      { S7_Templates := "SrcType := Real" } EQ_Contact(in1 := "MB_MFC_FLOAT_DB".FCounterLimit, in2 := "MB_MFC_FLOAT_DB".MFC401_VOL_SP)
      { S7_Templates := "SrcType := Real" } LT_Contact(in1 := "PT402_VAL", in2 := "PT402_HIGH")
      { S7_Templates := "SrcType := Real" } GE_Contact(in1 := "PT601_VAL", in2 := "PT401_CALC_50PRCT")
      wire#w9
      I_Contact( "S6_3" )
      wire#w10
      Coil( "S6_2" )
   END_RUNG
   RUNG wire#w8
      Contact( "S6_2" )
   END_RUNG wire#w9
   RUNG wire#w10
      Move(in := -1, out1 => "MB_MFC_FLOAT_DB"."STEP")
      Move(in := 0, out1 => "MB_MFC_INT_DB".MFC_Setpoint)
      Move(in := 40, out1 => "MB_MFC_INT_DB".START_STEP)   // Closes Valve
      S_Coil( "MB_MFC_INT_DB".LOAD_STEP )
   END_RUNG
   RUNG wire#w10
      S_Coil( "PV702_NC" )
   END_RUNG
   RUNG wire#powerrail
      Contact( #RUN )
      wire#w11
      Contact( "S6_2" )
      I_Contact( "PV702_NOT_OPEN_LS" )
      wire#w12
      { S7_Templates := "SrcType := SInt" } GE_Contact(in1 := "MB_MFC_INT_DB"."STEP", in2 := 2)
      { S7_Templates := "SrcType := UInt" } EQ_Contact(in1 := "MB_MFC_INT_DB".ControlMode, in2 := 0)
      { S7_Templates := "SrcType := UInt" } EQ_Contact(in1 := "MB_MFC_INT_DB".ValveOutput, in2 := 0)
      { S7_Templates := "SrcType := UInt" } EQ_Contact(in1 := "MB_MFC_INT_DB".Measure, in2 := 0)
      wire#w13
      I_Contact( "S6_3A" )
      wire#w14
      Coil( "S6_3" )
   END_RUNG
   RUNG wire#w12
      { S7_Templates := "SrcType := Real" } LE_Contact(in1 := "PT601_VAL", in2 := "PT901_VAL")
   END_RUNG wire#w13
   RUNG wire#w11
      Contact( "S6_3" )
   END_RUNG wire#w13
   RUNG wire#w14
      R_Coil( "PV702_NC" )
   END_RUNG
   RUNG wire#powerrail
      Contact( #RUN )
      wire#w15
      Contact( "S6_3" )
      I_Contact( "PV702_NOT_CLOSED_LS" )
      { S7_Templates := "SrcType := SInt" } GE_Contact(in1 := "MB_MFC_INT_DB"."STEP", in2 := 3)
      { S7_Templates := "SrcType := UInt" } EQ_Contact(in1 := "MB_MFC_INT_DB".CounterMode, in2 := 2)
      { S7_Templates := "SrcType := UInt" } EQ_Contact(in1 := "MB_MFC_INT_DB".CounterVal, in2 := 0)
      { S7_Templates := "SrcType := UInt" } EQ_Contact(in1 := "MB_MFC_INT_DB".ValveOutput, in2 := 0)
      { S7_Templates := "SrcType := UInt" } EQ_Contact(in1 := "MB_MFC_INT_DB".Measure, in2 := 0)
      I_Contact( #ALARM )
      wire#w16
      I_Contact( "S6_3B" )
      wire#w17
      Coil( "S6_3A" )
   END_RUNG
   RUNG wire#w15
      Contact( "S6_3A" )
   END_RUNG wire#w16
   RUNG wire#w17
      Move(in := -1, out1 => "MB_MFC_INT_DB"."STEP")
      Move(in := -1, out1 => "MB_MFC_FLOAT_DB"."STEP")
   END_RUNG
   RUNG wire#powerrail
      Contact( #RUN )
      wire#w18
      Contact( "S6_3A" )
      Contact( "IEC_Timer_S6_DB_1".Q )
      I_Contact( #ALARM )
      wire#w19
      I_Contact( "S6_4" )
      wire#w20
      Coil( "S6_3B" )
   END_RUNG
   RUNG wire#w18
      Contact( "S6_3B" )
   END_RUNG wire#w19
   RUNG wire#w20
      S_Coil( "PV701_NC" )
   END_RUNG
   RUNG wire#w20
      Move(in := "MB_MFC_FLOAT_DB".MFC401_FLOW_SP, out1 => "MB_MFC_FLOAT_DB".FLOW_SP)
      Move(in := 20, out1 => "MB_MFC_FLOAT_DB".START_STEP)
      S_Coil( "MB_MFC_FLOAT_DB".LOAD_STEP )
   END_RUNG
   RUNG wire#powerrail
      Contact( #RUN )
      wire#w21
      Contact( "S6_3B" )
      I_Contact( "PV701_NOT_OPEN_LS" )
      { S7_Templates := "SrcType := SInt" } EQ_Contact(in1 := "MB_MFC_FLOAT_DB"."STEP", in2 := 2)
      wire#w22
      I_Contact( "S6_5" )
      wire#w23
      Coil( "S6_4" )
   END_RUNG
   RUNG wire#w21
      Contact( "S6_4" )
   END_RUNG wire#w22
   RUNG wire#w23
      Move(in := -1, out1 => "MB_MFC_INT_DB"."STEP")
   END_RUNG
   RUNG wire#powerrail
      Contact( #RUN )
      wire#w24
      Contact( "S6_4" )
      wire#w25
      { S7_Templates := "SrcType := SInt" } GE_Contact(in1 := "MB_MFC_FLOAT_DB"."STEP", in2 := 1)
      { S7_Templates := "SrcType := Real" } GE_Contact(in1 := "MB_MFC_FLOAT_DB".FCounterVal, in2 := "MB_MFC_FLOAT_DB".COUNTER_LIMIT_SP)
      wire#w26
      I_Contact( "S6_6" )
      wire#w27
      Coil( "S6_5" )
   END_RUNG
   RUNG wire#w25
      { S7_Templates := "SrcType := Real" } GE_Contact(in1 := "PT901_VAL", in2 := "PT901_SP_H")
   END_RUNG wire#w26
   RUNG wire#w24
      Contact( "S6_5" )
   END_RUNG wire#w26
   RUNG wire#w27
      R_Coil( "PV401_NC" )
      R_Coil( "PV701_NC" )
   END_RUNG
   RUNG wire#w27
      Move(in := -1, out1 => "MB_MFC_FLOAT_DB"."STEP")
      Move(in := "MFC_601_MB_ADDR", out1 => "MB_MFC_INT_DB".MFC_ADDRESS)
      Move(in := 68, out1 => "MB_MFC_INT_DB".START_STEP)   // Purge Valve
      S_Coil( "MB_MFC_INT_DB".LOAD_STEP )
   END_RUNG
   RUNG wire#powerrail
      Contact( #RUN )
      wire#w28
      Contact( "S6_5" )
      I_Contact( "PV701_NOT_CLOSED_LS" )
      { S7_Templates := "SrcType := UInt" } EQ_Contact(in1 := "MB_MFC_INT_DB".ControlMode, in2 := 8)
      { S7_Templates := "SrcType := SInt" } EQ_Contact(in1 := "MB_MFC_INT_DB"."STEP", in2 := 4)
      wire#w29
      I_Contact( "S6_7" )
      wire#w30
      Coil( "S6_6" )
   END_RUNG
   RUNG wire#w28
      Contact( "S6_6" )
   END_RUNG wire#w29
   RUNG wire#w30
      S_Coil( "PV702_NC" )
   END_RUNG
   RUNG wire#w30
      Move(in := -1, out1 => "MB_MFC_INT_DB"."STEP")
   END_RUNG
   RUNG wire#powerrail
      Contact( #RUN )
      wire#w31
      Contact( "S6_6" )
      I_Contact( "PV702_NOT_OPEN_LS" )
      { S7_Templates := "SrcType := Real" } LE_Contact(in1 := "PT601_VAL", in2 := "PT601_ZERO")
      wire#w32
      I_Contact( "S6_8" )
      wire#w33
      Coil( "S6_7" )
   END_RUNG
   RUNG wire#w31
      Contact( "S6_7" )
   END_RUNG wire#w32
   RUNG wire#w33
      R_Coil( "PV602_NC" )
      R_Coil( "PV402_NC" )
   END_RUNG
   RUNG wire#w33
      R_Coil( "PV702_NC" )
   END_RUNG
   RUNG wire#w33
      Move(in := "MFC_601_MB_ADDR", out1 => "MB_MFC_INT_DB".MFC_ADDRESS)
      Move(in := "MB_VAL_CONTROL_MODE_BUS", out1 => "MB_MFC_INT_DB".MFC_MODE_SP)
      Move(in := 0, out1 => "MB_MFC_INT_DB".MFC_Setpoint)
      Move(in := 10, out1 => "MB_MFC_INT_DB".START_STEP)
      S_Coil( "MB_MFC_INT_DB".LOAD_STEP )
   END_RUNG
   RUNG wire#powerrail
      Contact( #RUN )
      wire#w34
      Contact( "S6_7" )
      I_Contact( "PV702_NOT_CLOSED_LS" )
      { S7_Templates := "SrcType := SInt" } EQ_Contact(in1 := "MB_MFC_INT_DB"."STEP", in2 := 4)
      { S7_Templates := "SrcType := UInt" } EQ_Contact(in1 := "MB_MFC_INT_DB".ControlMode, in2 := 0)
      Contact( "IEC_Timer_S6_DB_1".Q )
      wire#w35
      I_Contact( "S6_9" )
      wire#w36
      Coil( "S6_8" )
   END_RUNG
   RUNG wire#w34
      Contact( "S6_8" )
   END_RUNG wire#w35
   RUNG wire#w36
      R_Coil( "PV403_NO" )
   END_RUNG
   RUNG wire#w36
      { S7_GenerateENO := "TRUE" } Move(in := "PT901_VAL", out1 => "PT901_END_H")
   END_RUNG
   RUNG wire#w36
      Contact( "AlwaysFALSE" )
      Move(in := -1, out1 => "MB_MFC_INT_DB"."STEP")
      Move(in := -1, out1 => "MB_MFC_FLOAT_DB"."STEP")
   END_RUNG
   RUNG wire#powerrail
      Contact( #RUN )
      wire#w37
      Contact( "S6_8" )
      { S7_Templates := "SrcType := Real" } LE_Contact(in1 := "PT402_VAL", in2 := 0.0)
      wire#w38
      Coil( "S6_9" )
   END_RUNG
   RUNG wire#w37
      Contact( "S6_9" )
   END_RUNG wire#w38
   RUNG wire#w38
      Coil( #ENDED )
   END_RUNG
   // the same network as SCL:
   #_w1 := #RUN AND "AUTO_CYCLE" AND #RUN AND NOT "S6_M";   // rising edge of #RUN
   "S6_M" := #RUN;
   "S6_0" := ((((#RUN AND #START) OR #_w1) AND NOT #ALARM) OR (#RUN AND "S6_0")) AND NOT "S6_1";
   IF "S6_0" THEN
       "MB_MFC_FLOAT_DB".MFC_ADDRESS := "MFC_401_MB_ADDR";
       "MB_MFC_FLOAT_DB"."STEP" := -1;
       "MB_MFC_INT_DB".MFC_MODE_SP := "MB_VAL_CONTROL_MODE_BUS";
       "MB_MFC_INT_DB".START_STEP := 10;
       "MB_MFC_INT_DB".LOAD_STEP := TRUE;
       "MB_MFC_INT_DB".MFC_ADDRESS := "MFC_401_MB_ADDR";
       "GREEN_LIGHT" := FALSE;
       "YELLOW_LIGHT" := FALSE;
       "RED_ON" := TRUE;
   END_IF;
   "S6_1" := #RUN AND (("S6_0" AND "IEC_Timer_S6_DB_1".Q AND NOT #ALARM) OR "S6_1") AND NOT "S6_2";
   IF "S6_1" THEN
       "PV403_NO" := TRUE;
       "PV401_NC" := TRUE;
       "PV402_NC" := TRUE;
       "PV602_NC" := TRUE;
       "MB_MFC_INT_DB"."STEP" := -1;
       "MB_MFC_FLOAT_DB".FLOW_SP := 2.0;
       "MB_MFC_FLOAT_DB".START_STEP := 20;
       "MB_MFC_FLOAT_DB".LOAD_STEP := TRUE;
   END_IF;
   "S6_2" := #RUN AND (("S6_1" AND ("MB_MFC_FLOAT_DB"."STEP" >= 4) AND ("MB_MFC_FLOAT_DB".FCounterLimit = "MB_MFC_FLOAT_DB".MFC401_VOL_SP) AND ("PT402_VAL" < "PT402_HIGH") AND ("PT601_VAL" >= "PT401_CALC_50PRCT")) OR "S6_2") AND NOT "S6_3";
   IF "S6_2" THEN
       "MB_MFC_FLOAT_DB"."STEP" := -1;
       "MB_MFC_INT_DB".MFC_Setpoint := 0;
       "MB_MFC_INT_DB".START_STEP := 40;   // Closes Valve
       "MB_MFC_INT_DB".LOAD_STEP := TRUE;
       "PV702_NC" := TRUE;
   END_IF;
   "S6_3" := #RUN AND (("S6_2" AND NOT "PV702_NOT_OPEN_LS" AND ((("MB_MFC_INT_DB"."STEP" >= 2) AND ("MB_MFC_INT_DB".ControlMode = 0) AND ("MB_MFC_INT_DB".ValveOutput = 0) AND ("MB_MFC_INT_DB".Measure = 0)) OR ("PT601_VAL" <= "PT901_VAL"))) OR "S6_3") AND NOT "S6_3A";
   IF "S6_3" THEN "PV702_NC" := FALSE; END_IF;
   "S6_3A" := #RUN AND (("S6_3" AND NOT "PV702_NOT_CLOSED_LS" AND ("MB_MFC_INT_DB"."STEP" >= 3) AND ("MB_MFC_INT_DB".CounterMode = 2) AND ("MB_MFC_INT_DB".CounterVal = 0) AND ("MB_MFC_INT_DB".ValveOutput = 0) AND ("MB_MFC_INT_DB".Measure = 0) AND NOT #ALARM) OR "S6_3A") AND NOT "S6_3B";
   IF "S6_3A" THEN
       "MB_MFC_INT_DB"."STEP" := -1;
       "MB_MFC_FLOAT_DB"."STEP" := -1;
   END_IF;
   "S6_3B" := #RUN AND (("S6_3A" AND "IEC_Timer_S6_DB_1".Q AND NOT #ALARM) OR "S6_3B") AND NOT "S6_4";
   IF "S6_3B" THEN
       "PV701_NC" := TRUE;
       "MB_MFC_FLOAT_DB".FLOW_SP := "MB_MFC_FLOAT_DB".MFC401_FLOW_SP;
       "MB_MFC_FLOAT_DB".START_STEP := 20;
       "MB_MFC_FLOAT_DB".LOAD_STEP := TRUE;
   END_IF;
   "S6_4" := #RUN AND (("S6_3B" AND NOT "PV701_NOT_OPEN_LS" AND ("MB_MFC_FLOAT_DB"."STEP" = 2)) OR "S6_4") AND NOT "S6_5";
   IF "S6_4" THEN "MB_MFC_INT_DB"."STEP" := -1; END_IF;
   "S6_5" := #RUN AND (("S6_4" AND ((("MB_MFC_FLOAT_DB"."STEP" >= 1) AND ("MB_MFC_FLOAT_DB".FCounterVal >= "MB_MFC_FLOAT_DB".COUNTER_LIMIT_SP)) OR ("PT901_VAL" >= "PT901_SP_H"))) OR "S6_5") AND NOT "S6_6";
   IF "S6_5" THEN
       "PV401_NC" := FALSE;
       "PV701_NC" := FALSE;
       "MB_MFC_FLOAT_DB"."STEP" := -1;
       "MB_MFC_INT_DB".MFC_ADDRESS := "MFC_601_MB_ADDR";
       "MB_MFC_INT_DB".START_STEP := 68;   // Purge Valve
       "MB_MFC_INT_DB".LOAD_STEP := TRUE;
   END_IF;
   "S6_6" := #RUN AND (("S6_5" AND NOT "PV701_NOT_CLOSED_LS" AND ("MB_MFC_INT_DB".ControlMode = 8) AND ("MB_MFC_INT_DB"."STEP" = 4)) OR "S6_6") AND NOT "S6_7";
   IF "S6_6" THEN
       "PV702_NC" := TRUE;
       "MB_MFC_INT_DB"."STEP" := -1;
   END_IF;
   "S6_7" := #RUN AND (("S6_6" AND NOT "PV702_NOT_OPEN_LS" AND ("PT601_VAL" <= "PT601_ZERO")) OR "S6_7") AND NOT "S6_8";
   IF "S6_7" THEN
       "PV602_NC" := FALSE;
       "PV402_NC" := FALSE;
       "PV702_NC" := FALSE;
       "MB_MFC_INT_DB".MFC_ADDRESS := "MFC_601_MB_ADDR";
       "MB_MFC_INT_DB".MFC_MODE_SP := "MB_VAL_CONTROL_MODE_BUS";
       "MB_MFC_INT_DB".MFC_Setpoint := 0;
       "MB_MFC_INT_DB".START_STEP := 10;
       "MB_MFC_INT_DB".LOAD_STEP := TRUE;
   END_IF;
   "S6_8" := #RUN AND (("S6_7" AND NOT "PV702_NOT_CLOSED_LS" AND ("MB_MFC_INT_DB"."STEP" = 4) AND ("MB_MFC_INT_DB".ControlMode = 0) AND "IEC_Timer_S6_DB_1".Q) OR "S6_8") AND NOT "S6_9";
   IF "S6_8" THEN
       "PV403_NO" := FALSE;
       "PT901_END_H" := "PT901_VAL";
   END_IF;
   IF "S6_8" AND "AlwaysFALSE" THEN
       "MB_MFC_INT_DB"."STEP" := -1;
       "MB_MFC_FLOAT_DB"."STEP" := -1;
   END_IF;
   "S6_9" := #RUN AND (("S6_8" AND ("PT402_VAL" <= 0.0)) OR "S6_9");
   #ENDED := "S6_9";
END_REGION

REGION Network 4
   // Timers
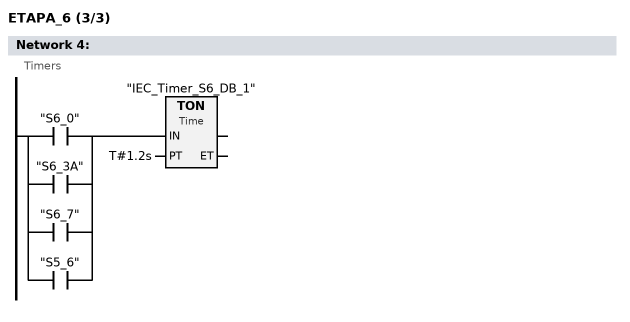
   "IEC_Timer_S6_DB_1".TON(IN := "S6_0" OR "S6_3A" OR "S6_7" OR "S5_6", PT := T#1.2s);
END_REGION
END_FUNCTION

FUNCTION "ETAPA_7" : Void   // FC8, LAD
TITLE = CICLO de INJECÇÃO - injecção de Hélio 2
{ S7_Optimized_Access := 'FALSE' }
VERSION : 0.1
   VAR_TEMP   // added for the SCL form of the ladder/FBD networks
      _w1 : Bool;
   END_VAR
BEGIN

REGION Network 1
   // PT Alarm  Set Points
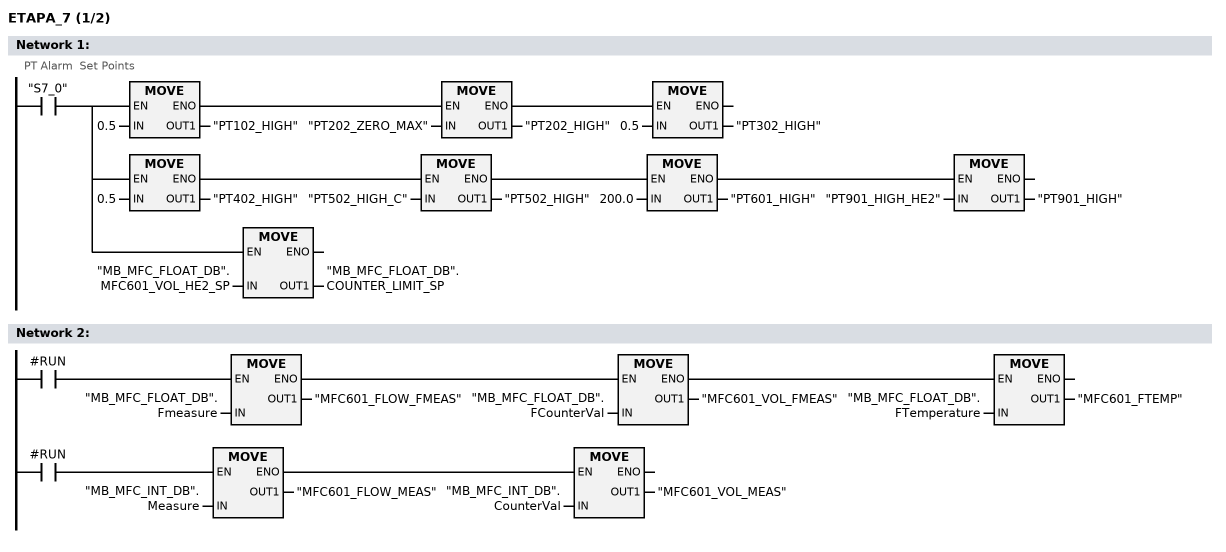
   RUNG wire#powerrail
      Contact( "S7_0" )
      wire#w1
      { S7_GenerateENO := "TRUE" } Move(in := 0.5, out1 => "PT102_HIGH")
      { S7_GenerateENO := "TRUE" } Move(in := "PT202_ZERO_MAX", out1 => "PT202_HIGH")
      { S7_GenerateENO := "TRUE" } Move(in := 0.5, out1 => "PT302_HIGH")
   END_RUNG
   RUNG wire#w1
      { S7_GenerateENO := "TRUE" } Move(in := 0.5, out1 => "PT402_HIGH")
      { S7_GenerateENO := "TRUE" } Move(in := "PT502_HIGH_C", out1 => "PT502_HIGH")
      { S7_GenerateENO := "TRUE" } Move(in := 200.0, out1 => "PT601_HIGH")
      { S7_GenerateENO := "TRUE" } Move(in := "PT901_HIGH_HE2", out1 => "PT901_HIGH")
   END_RUNG
   RUNG wire#w1
      Move(in := "MB_MFC_FLOAT_DB".MFC601_VOL_HE2_SP, out1 => "MB_MFC_FLOAT_DB".COUNTER_LIMIT_SP)
   END_RUNG
   // the same network as SCL:
   // ENO of a box is taken as its EN; it also drops when the box reports an error
   IF "S7_0" THEN
       "PT102_HIGH" := 0.5;
       "PT202_HIGH" := "PT202_ZERO_MAX";
       "PT302_HIGH" := 0.5;
       "PT402_HIGH" := 0.5;
       "PT502_HIGH" := "PT502_HIGH_C";
       "PT601_HIGH" := 200.0;
       "PT901_HIGH" := "PT901_HIGH_HE2";
       "MB_MFC_FLOAT_DB".COUNTER_LIMIT_SP := "MB_MFC_FLOAT_DB".MFC601_VOL_HE2_SP;
   END_IF;
END_REGION

REGION Network 2
   RUNG wire#powerrail
      Contact( #RUN )
      { S7_GenerateENO := "TRUE" } Move(in := "MB_MFC_FLOAT_DB".Fmeasure, out1 => "MFC601_FLOW_FMEAS")
      { S7_GenerateENO := "TRUE" } Move(in := "MB_MFC_FLOAT_DB".FCounterVal, out1 => "MFC601_VOL_FMEAS")
      { S7_GenerateENO := "TRUE" } Move(in := "MB_MFC_FLOAT_DB".FTemperature, out1 => "MFC601_FTEMP")
   END_RUNG
   RUNG wire#powerrail
      Contact( #RUN )
      { S7_GenerateENO := "TRUE" } Move(in := "MB_MFC_INT_DB".Measure, out1 => "MFC601_FLOW_MEAS")
      { S7_GenerateENO := "TRUE" } Move(in := "MB_MFC_INT_DB".CounterVal, out1 => "MFC601_VOL_MEAS")
   END_RUNG
   // the same network as SCL:
   // ENO of a box is taken as its EN; it also drops when the box reports an error
   IF #RUN THEN
       "MFC601_FLOW_FMEAS" := "MB_MFC_FLOAT_DB".Fmeasure;
       "MFC601_VOL_FMEAS" := "MB_MFC_FLOAT_DB".FCounterVal;
       "MFC601_FTEMP" := "MB_MFC_FLOAT_DB".FTemperature;
       "MFC601_FLOW_MEAS" := "MB_MFC_INT_DB".Measure;
       "MFC601_VOL_MEAS" := "MB_MFC_INT_DB".CounterVal;
   END_IF;
END_REGION

REGION Network 3
   // Logica do ciclo 6
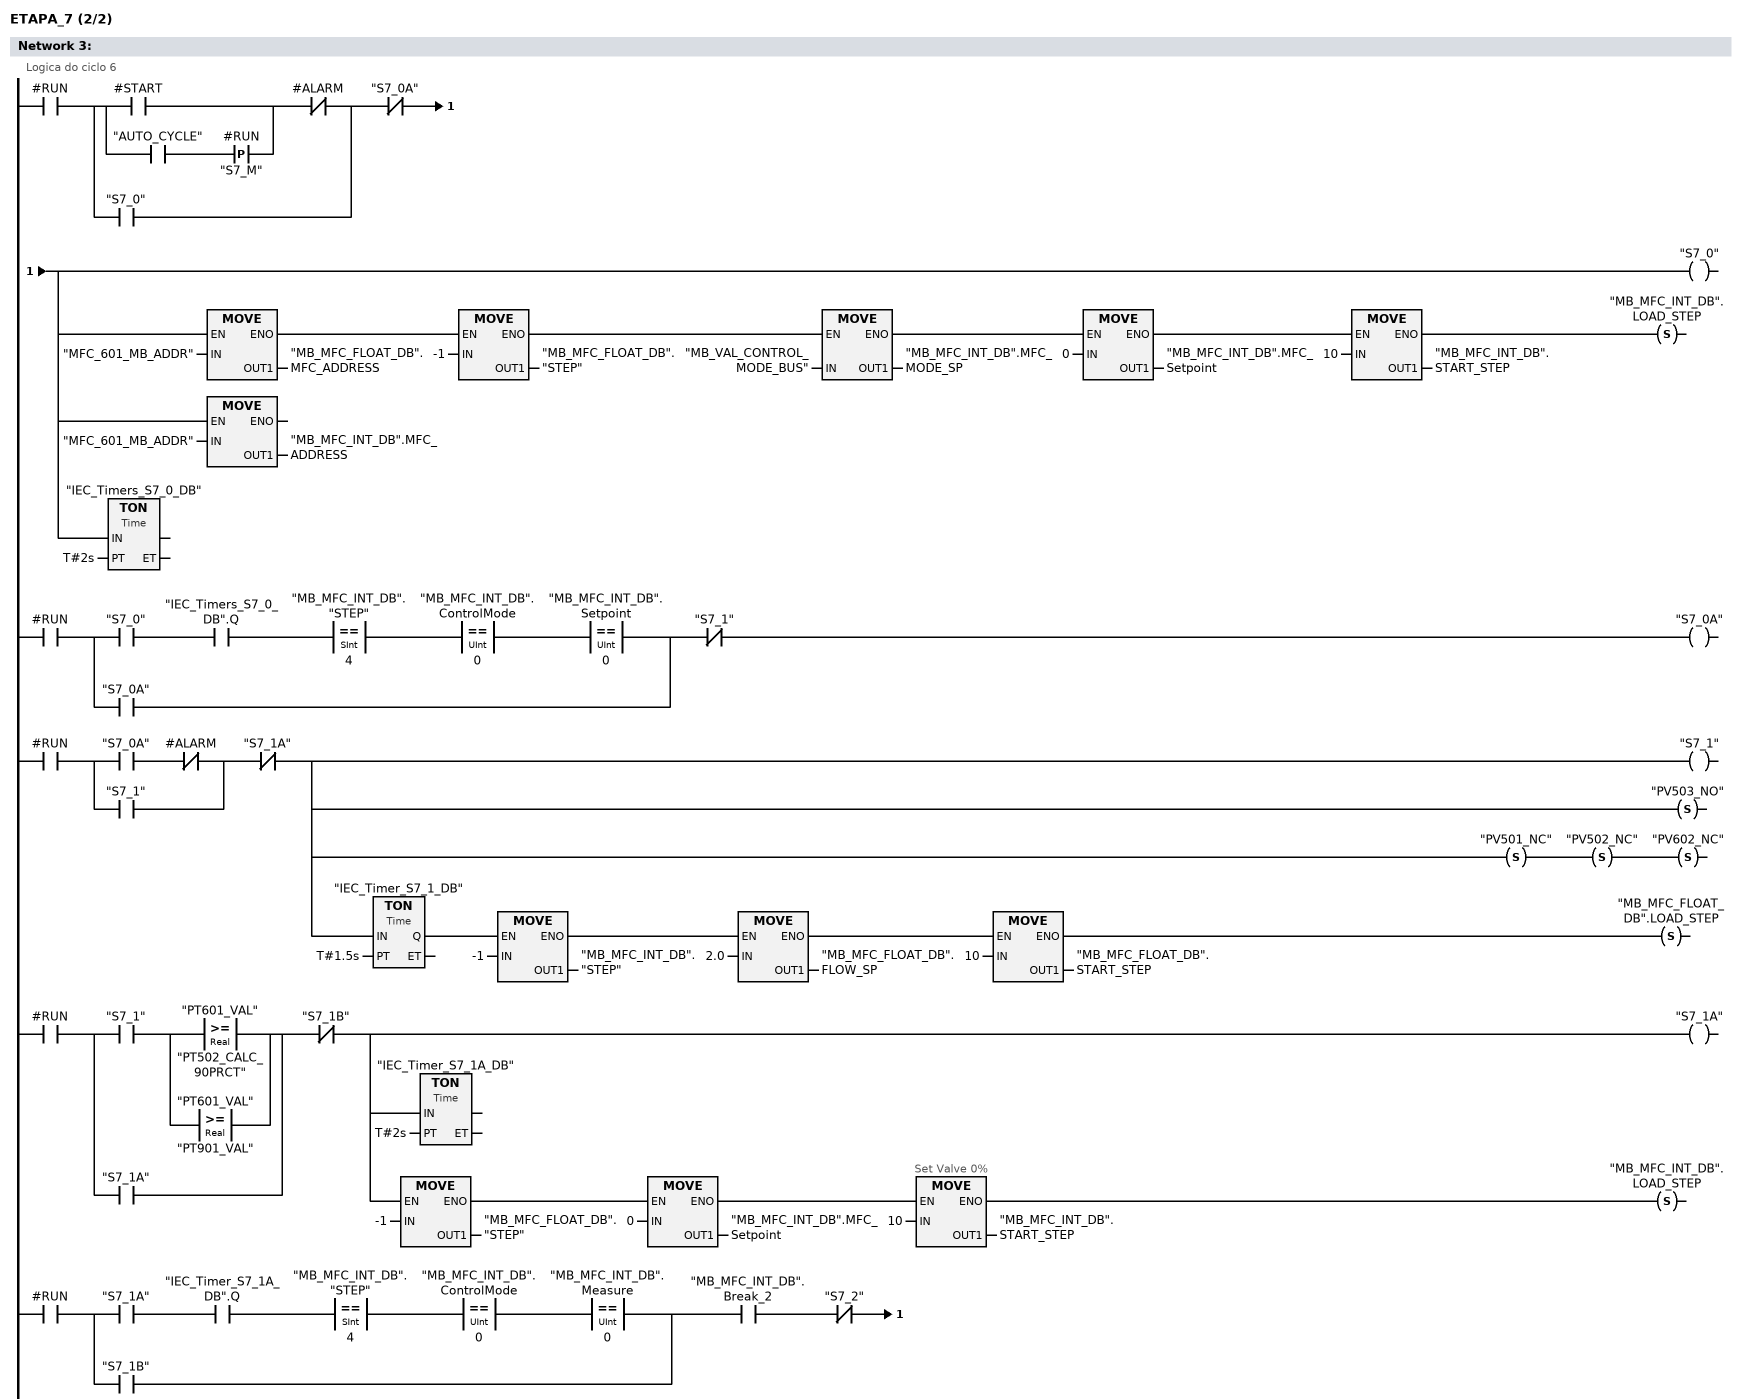
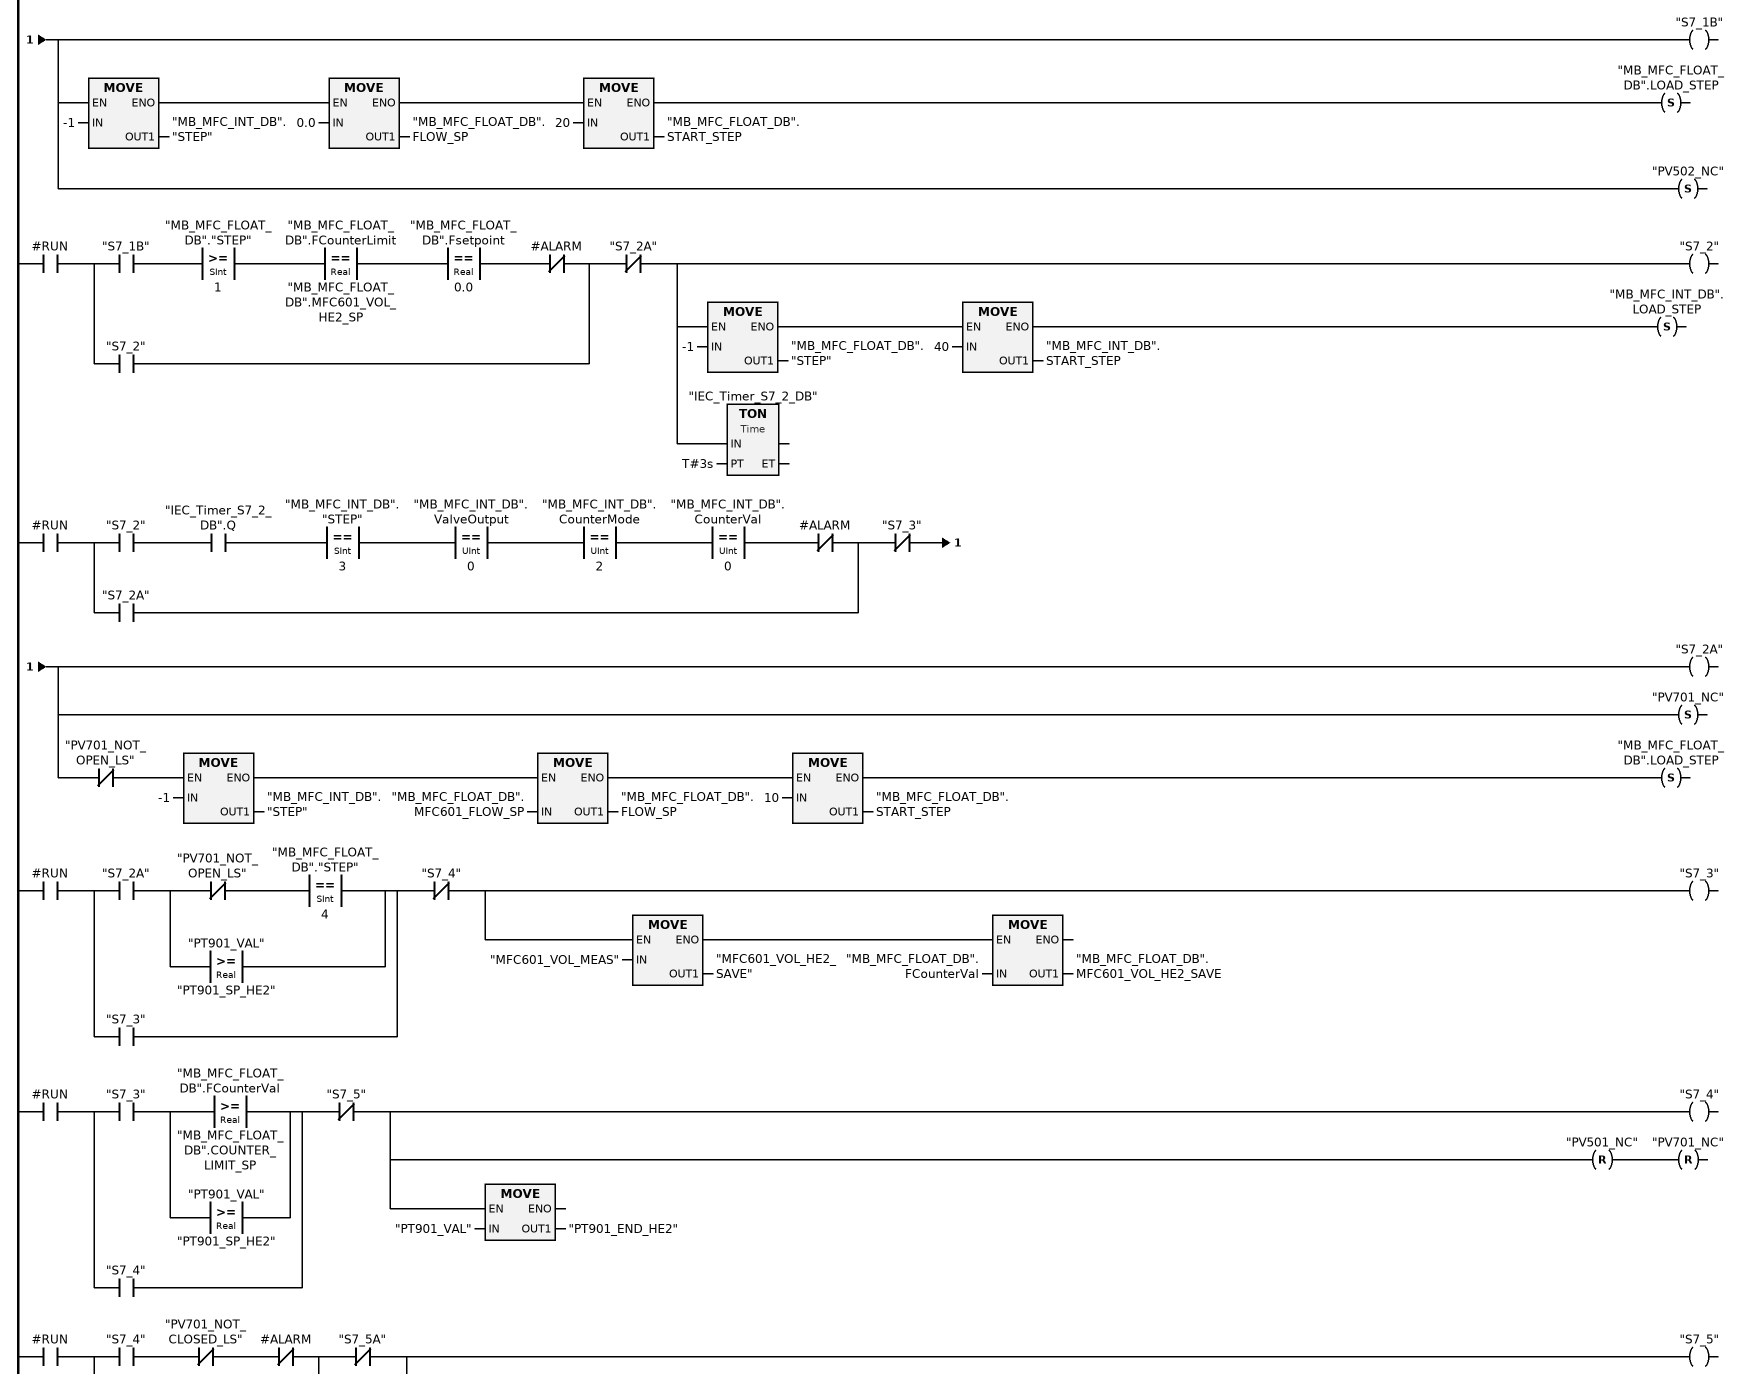
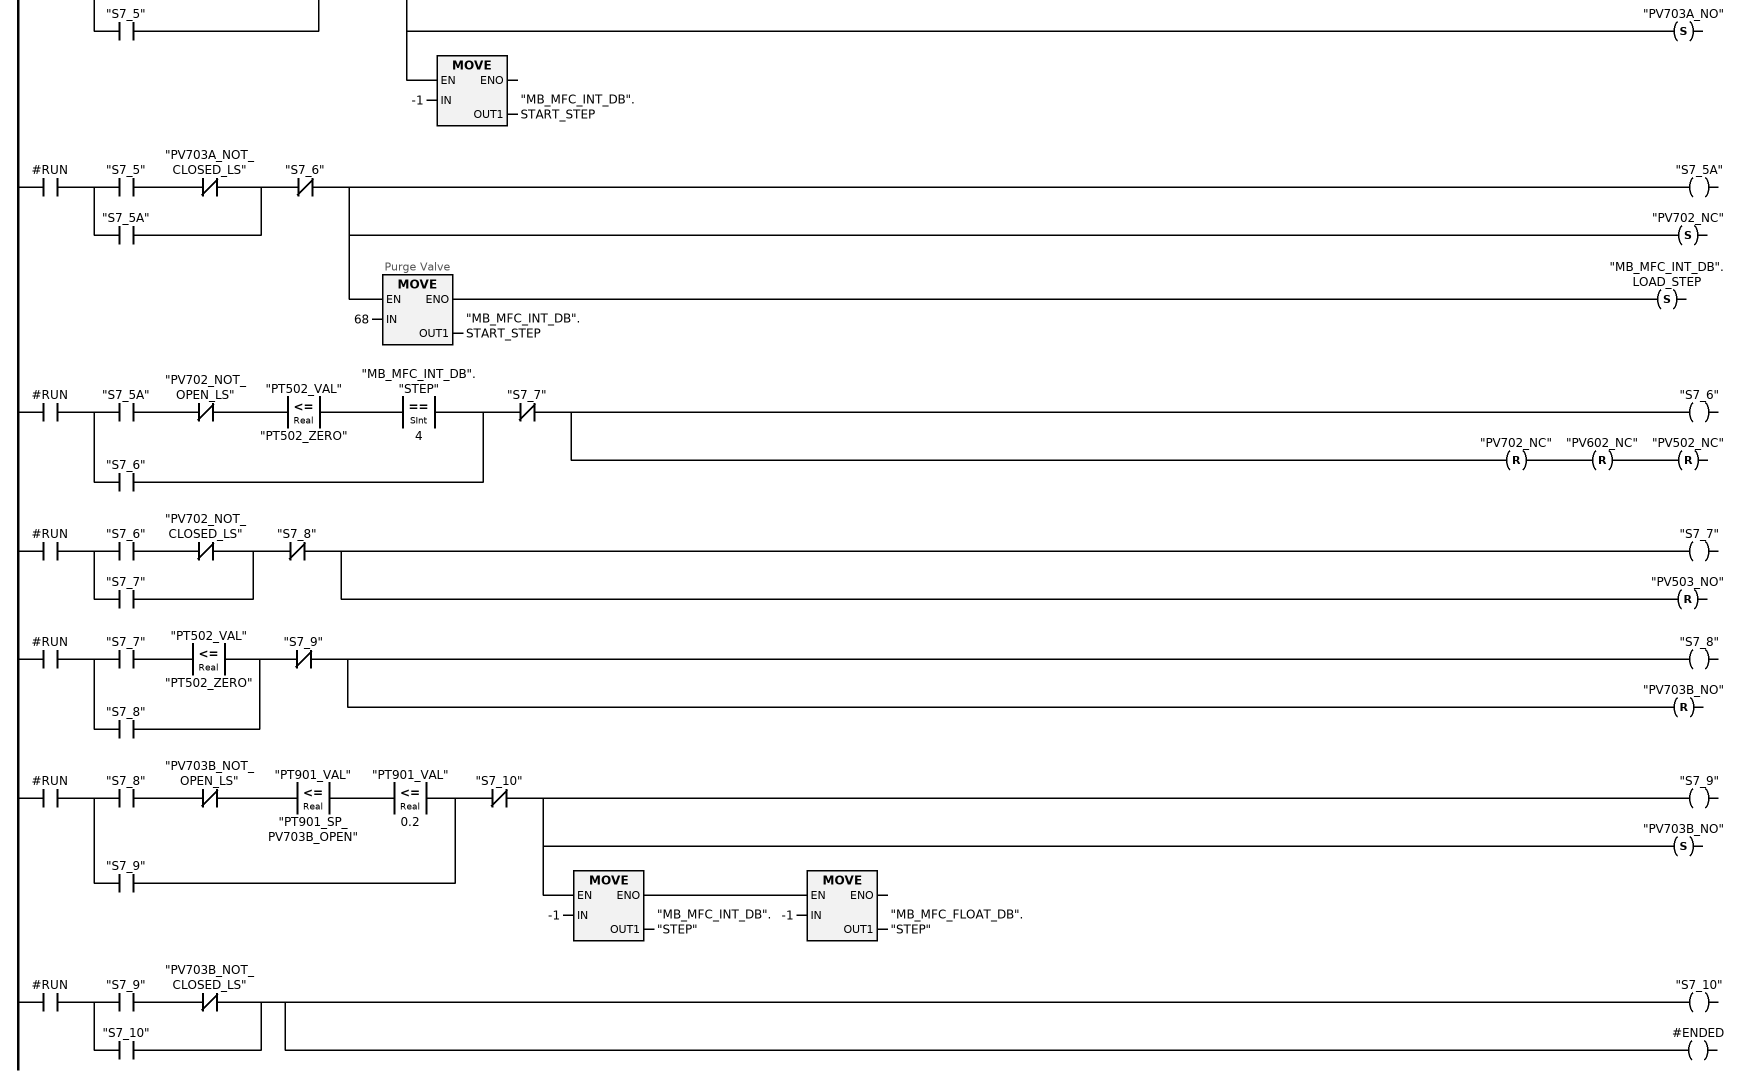
   #_w1 := #RUN AND "AUTO_CYCLE" AND #RUN AND NOT "S7_M";   // rising edge of #RUN
   "S7_M" := #RUN;
   "S7_0" := ((((#RUN AND #START) OR #_w1) AND NOT #ALARM) OR (#RUN AND "S7_0")) AND NOT "S7_0A";
   IF "S7_0" THEN
       "MB_MFC_FLOAT_DB".MFC_ADDRESS := "MFC_601_MB_ADDR";
       "MB_MFC_FLOAT_DB"."STEP" := -1;
       "MB_MFC_INT_DB".MFC_MODE_SP := "MB_VAL_CONTROL_MODE_BUS";
       "MB_MFC_INT_DB".MFC_Setpoint := 0;
       "MB_MFC_INT_DB".START_STEP := 10;
       "MB_MFC_INT_DB".LOAD_STEP := TRUE;
       "MB_MFC_INT_DB".MFC_ADDRESS := "MFC_601_MB_ADDR";
   END_IF;
   "IEC_Timers_S7_0_DB".TON(IN := "S7_0", PT := T#2s);
   "S7_0A" := #RUN AND (("S7_0" AND "IEC_Timers_S7_0_DB".Q AND ("MB_MFC_INT_DB"."STEP" = 4) AND ("MB_MFC_INT_DB".ControlMode = 0) AND ("MB_MFC_INT_DB".Setpoint = 0)) OR "S7_0A") AND NOT "S7_1";
   "S7_1" := #RUN AND (("S7_0A" AND NOT #ALARM) OR "S7_1") AND NOT "S7_1A";
   IF "S7_1" THEN
       "PV503_NO" := TRUE;
       "PV501_NC" := TRUE;
       "PV502_NC" := TRUE;
       "PV602_NC" := TRUE;
   END_IF;
   "IEC_Timer_S7_1_DB".TON(IN := "S7_1", PT := T#1.5s);
   IF "IEC_Timer_S7_1_DB".Q THEN
       "MB_MFC_INT_DB"."STEP" := -1;
       "MB_MFC_FLOAT_DB".FLOW_SP := 2.0;
       "MB_MFC_FLOAT_DB".START_STEP := 10;
       "MB_MFC_FLOAT_DB".LOAD_STEP := TRUE;
   END_IF;
   "S7_1A" := #RUN AND (("S7_1" AND (("PT601_VAL" >= "PT502_CALC_90PRCT") OR ("PT601_VAL" >= "PT901_VAL"))) OR "S7_1A") AND NOT "S7_1B";
   "IEC_Timer_S7_1A_DB".TON(IN := "S7_1A", PT := T#2s);
   IF "S7_1A" THEN
       "MB_MFC_FLOAT_DB"."STEP" := -1;
       "MB_MFC_INT_DB".MFC_Setpoint := 0;
       "MB_MFC_INT_DB".START_STEP := 10;   // Set Valve 0%
       "MB_MFC_INT_DB".LOAD_STEP := TRUE;
   END_IF;
   "S7_1B" := #RUN AND (("S7_1A" AND "IEC_Timer_S7_1A_DB".Q AND ("MB_MFC_INT_DB"."STEP" = 4) AND ("MB_MFC_INT_DB".ControlMode = 0) AND ("MB_MFC_INT_DB".Measure = 0)) OR "S7_1B") AND "MB_MFC_INT_DB".Break_2 AND NOT "S7_2";
   IF "S7_1B" THEN
       "MB_MFC_INT_DB"."STEP" := -1;
       "MB_MFC_FLOAT_DB".FLOW_SP := 0.0;
       "MB_MFC_FLOAT_DB".START_STEP := 20;
       "MB_MFC_FLOAT_DB".LOAD_STEP := TRUE;
       "PV502_NC" := TRUE;
   END_IF;
   "S7_2" := #RUN AND (("S7_1B" AND ("MB_MFC_FLOAT_DB"."STEP" >= 1) AND ("MB_MFC_FLOAT_DB".FCounterLimit = "MB_MFC_FLOAT_DB".MFC601_VOL_HE2_SP) AND ("MB_MFC_FLOAT_DB".Fsetpoint = 0.0) AND NOT #ALARM) OR "S7_2") AND NOT "S7_2A";
   IF "S7_2" THEN
       "MB_MFC_FLOAT_DB"."STEP" := -1;
       "MB_MFC_INT_DB".START_STEP := 40;
       "MB_MFC_INT_DB".LOAD_STEP := TRUE;
   END_IF;
   "IEC_Timer_S7_2_DB".TON(IN := "S7_2", PT := T#3s);
   "S7_2A" := #RUN AND (("S7_2" AND "IEC_Timer_S7_2_DB".Q AND ("MB_MFC_INT_DB"."STEP" = 3) AND ("MB_MFC_INT_DB".ValveOutput = 0) AND ("MB_MFC_INT_DB".CounterMode = 2) AND ("MB_MFC_INT_DB".CounterVal = 0) AND NOT #ALARM) OR "S7_2A") AND NOT "S7_3";
   IF "S7_2A" THEN "PV701_NC" := TRUE; END_IF;
   IF "S7_2A" AND NOT "PV701_NOT_OPEN_LS" THEN
       "MB_MFC_INT_DB"."STEP" := -1;
       "MB_MFC_FLOAT_DB".FLOW_SP := "MB_MFC_FLOAT_DB".MFC601_FLOW_SP;
       "MB_MFC_FLOAT_DB".START_STEP := 10;
       "MB_MFC_FLOAT_DB".LOAD_STEP := TRUE;
   END_IF;
   "S7_3" := #RUN AND (("S7_2A" AND ((NOT "PV701_NOT_OPEN_LS" AND ("MB_MFC_FLOAT_DB"."STEP" = 4)) OR ("PT901_VAL" >= "PT901_SP_HE2"))) OR "S7_3") AND NOT "S7_4";
   IF "S7_3" THEN
       "MFC601_VOL_HE2_SAVE" := "MFC601_VOL_MEAS";
       "MB_MFC_FLOAT_DB".MFC601_VOL_HE2_SAVE := "MB_MFC_FLOAT_DB".FCounterVal;
   END_IF;
   "S7_4" := #RUN AND (("S7_3" AND (("MB_MFC_FLOAT_DB".FCounterVal >= "MB_MFC_FLOAT_DB".COUNTER_LIMIT_SP) OR ("PT901_VAL" >= "PT901_SP_HE2"))) OR "S7_4") AND NOT "S7_5";
   IF "S7_4" THEN
       "PV501_NC" := FALSE;
       "PV701_NC" := FALSE;
       "PT901_END_HE2" := "PT901_VAL";
   END_IF;
   "S7_5" := #RUN AND (("S7_4" AND NOT "PV701_NOT_CLOSED_LS" AND NOT #ALARM) OR "S7_5") AND NOT "S7_5A";
   IF "S7_5" THEN
       "PV703A_NO" := TRUE;
       "MB_MFC_INT_DB".START_STEP := -1;
   END_IF;
   "S7_5A" := #RUN AND (("S7_5" AND NOT "PV703A_NOT_CLOSED_LS") OR "S7_5A") AND NOT "S7_6";
   IF "S7_5A" THEN
       "PV702_NC" := TRUE;
       "MB_MFC_INT_DB".START_STEP := 68;   // Purge Valve
       "MB_MFC_INT_DB".LOAD_STEP := TRUE;
   END_IF;
   "S7_6" := #RUN AND (("S7_5A" AND NOT "PV702_NOT_OPEN_LS" AND ("PT502_VAL" <= "PT502_ZERO") AND ("MB_MFC_INT_DB"."STEP" = 4)) OR "S7_6") AND NOT "S7_7";
   IF "S7_6" THEN
       "PV702_NC" := FALSE;
       "PV602_NC" := FALSE;
       "PV502_NC" := FALSE;
   END_IF;
   "S7_7" := #RUN AND (("S7_6" AND NOT "PV702_NOT_CLOSED_LS") OR "S7_7") AND NOT "S7_8";
   IF "S7_7" THEN "PV503_NO" := FALSE; END_IF;
   "S7_8" := #RUN AND (("S7_7" AND ("PT502_VAL" <= "PT502_ZERO")) OR "S7_8") AND NOT "S7_9";
   IF "S7_8" THEN "PV703B_NO" := FALSE; END_IF;
   "S7_9" := #RUN AND (("S7_8" AND NOT "PV703B_NOT_OPEN_LS" AND ("PT901_VAL" <= "PT901_SP_PV703B_OPEN") AND ("PT901_VAL" <= 0.2)) OR "S7_9") AND NOT "S7_10";
   IF "S7_9" THEN
       "PV703B_NO" := TRUE;
       "MB_MFC_INT_DB"."STEP" := -1;
       "MB_MFC_FLOAT_DB"."STEP" := -1;
   END_IF;
   "S7_10" := #RUN AND (("S7_9" AND NOT "PV703B_NOT_CLOSED_LS") OR "S7_10");
   #ENDED := "S7_10";
END_REGION
END_FUNCTION

FUNCTION "ETAPA_8" : Void   // FC9, LAD
{ S7_Optimized_Access := 'FALSE' }
VERSION : 0.1
BEGIN
END_FUNCTION

FUNCTION "TESTS" : Void   // FC10, LAD
{ S7_Optimized_Access := 'FALSE' }
VERSION : 0.1
   VAR_TEMP   // added for the SCL form of the ladder/FBD networks
      _w1 : Bool;
   END_VAR
BEGIN

REGION Network 1
   // ALARM Settings
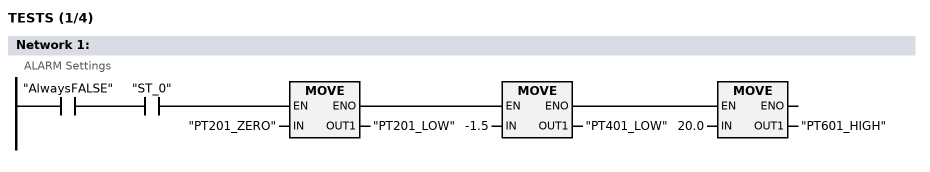
   RUNG wire#powerrail
      Contact( "AlwaysFALSE" )
      Contact( "ST_0" )
      { S7_GenerateENO := "TRUE" } Move(in := "PT201_ZERO", out1 => "PT201_LOW")
      { S7_GenerateENO := "TRUE" } Move(in := -1.5, out1 => "PT401_LOW")
      { S7_GenerateENO := "TRUE" } Move(in := 20.0, out1 => "PT601_HIGH")
   END_RUNG
   // the same network as SCL:
   // ENO of a box is taken as its EN; it also drops when the box reports an error
   IF "AlwaysFALSE" AND "ST_0" THEN
       "PT201_LOW" := "PT201_ZERO";
       "PT401_LOW" := -1.5;
       "PT601_HIGH" := 20.0;
   END_IF;
END_REGION

REGION Network 2: Pneumatic Tests
   // Test Pneumatic System (Test #1-#6)
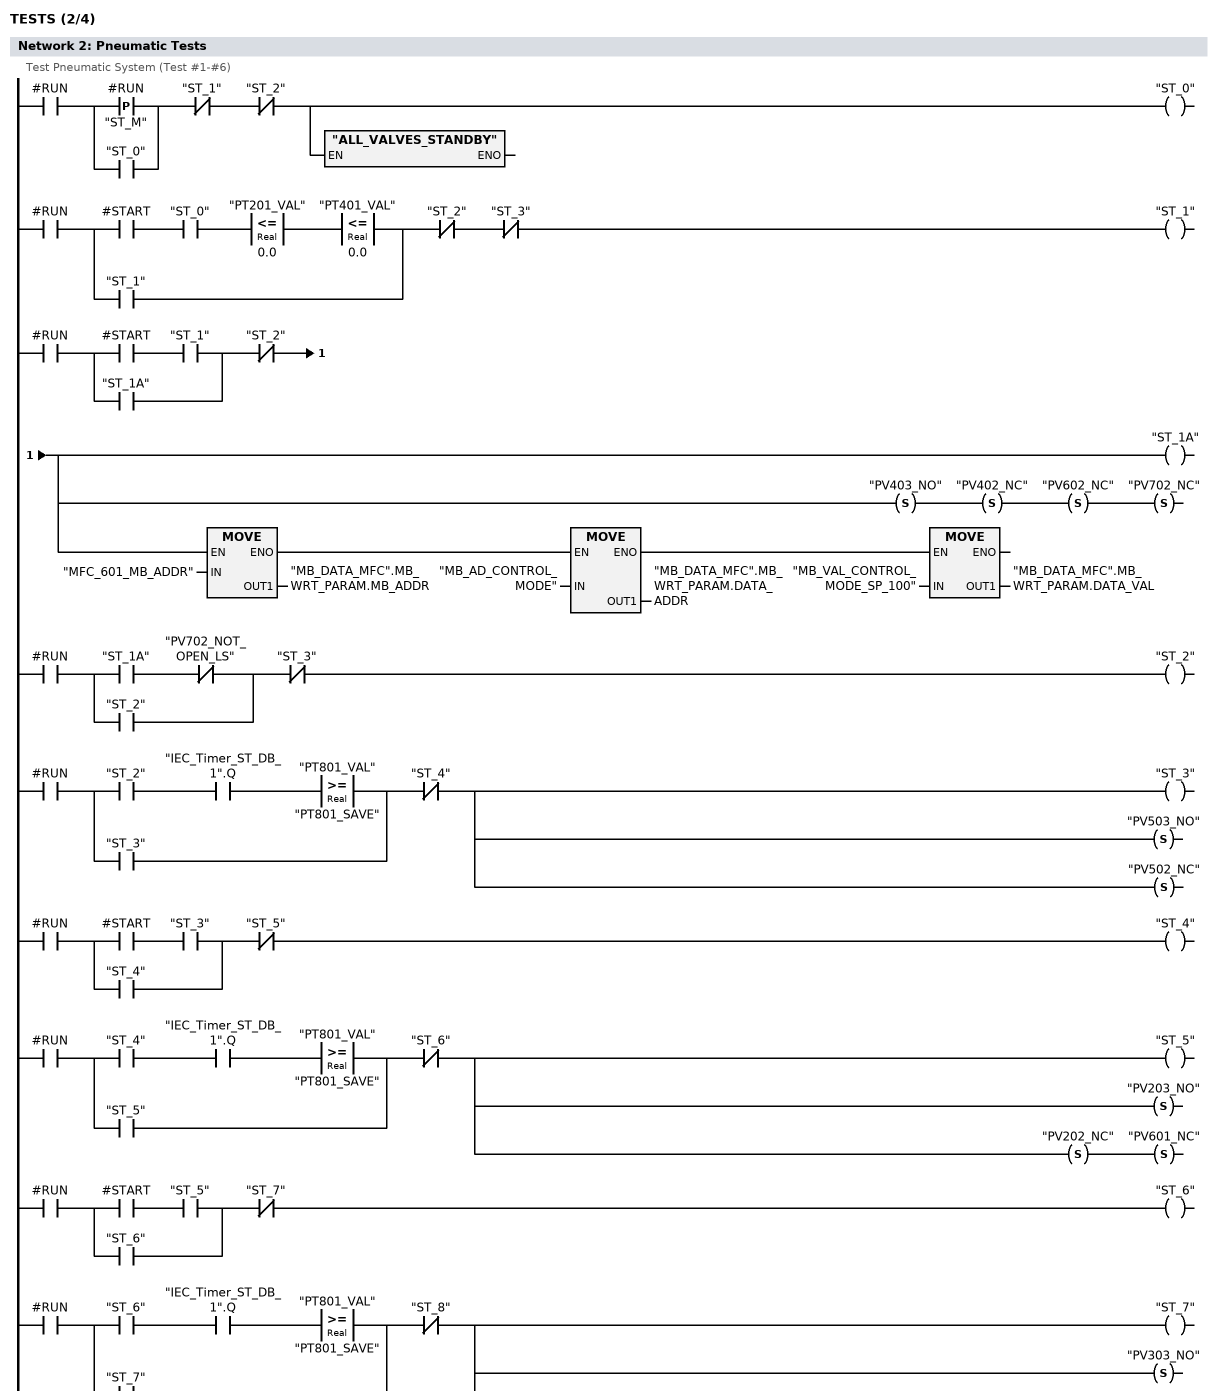
